// TIA Portal project "1215C_BREAKOUT_BOARD" (V19) (continued)
REGION Network 3
   RUNG wire#powerrail
      "FC10029_Custom_LGF_DTLtoString"(inDTL := "DB002-DateTime".LOCAL_DTL, format := 1, Ret_Val => "DB002-DateTime".DTLtoString_Ret, outDate_YY => "DB002-DateTime".sCustomDate_YY, outDate_MM => "DB002-DateTime".sCustomDate_MM, outDate_DD => "DB002-DateTime".sCustomDate_DD, outTime_HH => "DB002-DateTime".sCustomTime_HH, outTime_MM => "DB002-DateTime".sCustomTime_MM)
      "FC10030_Custom_DateTime_Format"(LOCAL_DTL := "DB002-DateTime".LOCAL_DTL, sCustomDate_YY := "DB002-DateTime".sCustomDate_YY, sCustomDate_MM := "DB002-DateTime".sCustomDate_MM, sCustomDate_DD := "DB002-DateTime".sCustomDate_DD, sCustomTime_HH := "DB002-DateTime".sCustomTime_HH, sCustomTime_MM := "DB002-DateTime".sCustomTime_MM, sCustomDate_DDMMYY := "DB002-DateTime".sCustomDate_DDMMYY, sCustomTime_HHMM := "DB002-DateTime".sCustomTime_HHMM)
   END_RUNG
   // the same network as SCL:
   "DB002-DateTime".DTLtoString_Ret := "FC10029_Custom_LGF_DTLtoString"(inDTL := "DB002-DateTime".LOCAL_DTL,
                           format := 1,
                           outDate_YY => "DB002-DateTime".sCustomDate_YY,
                           outDate_MM => "DB002-DateTime".sCustomDate_MM,
                           outDate_DD => "DB002-DateTime".sCustomDate_DD,
                           outTime_HH => "DB002-DateTime".sCustomTime_HH,
                           outTime_MM => "DB002-DateTime".sCustomTime_MM,
                           ENO => #_w1);
   IF #_w1 THEN
       "FC10030_Custom_DateTime_Format"(LOCAL_DTL := "DB002-DateTime".LOCAL_DTL,
                               sCustomDate_YY := "DB002-DateTime".sCustomDate_YY,
                               sCustomDate_MM := "DB002-DateTime".sCustomDate_MM,
                               sCustomDate_DD := "DB002-DateTime".sCustomDate_DD,
                               sCustomTime_HH := "DB002-DateTime".sCustomTime_HH,
                               sCustomTime_MM := "DB002-DateTime".sCustomTime_MM,
                               sCustomDate_DDMMYY := "DB002-DateTime".sCustomDate_DDMMYY,
                               sCustomTime_HHMM := "DB002-DateTime".sCustomTime_HHMM);
   END_IF;
END_REGION
END_FUNCTION

FUNCTION "FC10029_Custom_LGF_DTLtoString" : String   // FC10029, SCL
{ S7_Optimized_Access := 'TRUE' }
VERSION : 0.1
   VAR_INPUT
      inDTL : DTL;   // Date as DTL tag
      format : Bool;   // 1 = traditional, 0 = international
   END_VAR
   VAR_OUTPUT
      outDate_YY : String;   // Custom Date Output (YY)
      outDate_MM : String;   // Custom Date Output (MM)
      outDate_DD : String;   // Custom Date Output (DD)
      outTime_HH : String;   // Custom Time Output (HH)
      outTime_MM : String;   // Custom Time Output (MM)
   END_VAR
   VAR_TEMP
      tempString : String;   // -
      tempSepTime : Char;   // -
      tempPosYear : USInt;   // -
      tempPosMonth : USInt;   // -
      tempPosDay : USInt;   // -
      tempPosHour : USInt;   // -
      tempPosMinute : USInt;   // -
      tempPosSepYearMonth : USInt;   // -
      tempPosSepMonthDay : USInt;   // -
      tempPosSepHourMinute : USInt;   // -
   END_VAR
   // Ret_Val : Date as String tag
BEGIN
   //=============================================================================
   // Siemens AG
   // (c)Copyright 2017
   //-----------------------------------------------------------------------------
   // Library:       LGF (Library General Functions)
   // Tested with:   CPU1212C DC/DC/DC FW:V4.2
   // Engineering:   TIA Portal V14 Update 1
   // Restrictions:  -
   // Requirements:  PLC (S7-1200 / S7-1500)
   // Functionality: This function converts DTL into a string.  (EDITED)
   //-----------------------------------------------------------------------------
   // Change log table:
   // Version  Date        In charge / Changes applied
   // 01.00.00 15.06.2016  Siemens Industry Online Support
   //                      First released version
   // 01.00.01 02.01.2017  Siemens Industry Online Support
   //                      Upgrade: TIA Portal V14 Update 1
   // 01.00.02 17.08.2018  Siemens Industry Online Support
   //                      Upgrade: TIA V15 Update 2
   //=============================================================================


   // Initialization
   #tempString := '';
   #tempSepTime := ':';


   // Set format parameters for output string
   IF NOT #format
   THEN                                          // International ISO 8601
       #tempPosYear := 1;                          // DTL  | Y| Y| Y| Y| -| M| M| -| D| D|  | H| H| :| M| M|
       #tempPosMonth := 6;                         // -----|--|--|--|--|--|--|--|--|--|--|--|--|--|--|--|--|
       #tempPosDay := 9;                           // Pos  | 1| 2| 3| 4| 5| 6| 7| 8| 9|10|11|12|13|14|15|16|
       #tempPosHour := 12;
       #tempPosMinute := 15;
       #tempPosSepYearMonth := 5;
       #tempPosSepMonthDay := 8;
       #tempPosSepHourMinute := 14;
   ELSE                                          // Traditional (EU)
       #tempPosYear := 7;                          // DTL  | D| D| -| M| M| -| Y| Y| Y| Y|  | H| H| :| M| M|
       #tempPosMonth := 4;                         // -----|--|--|--|--|--|--|--|--|--|--|--|--|--|--|--|--|
       #tempPosDay := 1;                           // Pos  | 1| 2| 3| 4| 5| 6| 7| 8| 9|10|11|12|13|14|15|16|
       #tempPosHour := 12;
       #tempPosMinute := 15;
       #tempPosSepYearMonth := 6;
       #tempPosSepMonthDay := 3;
       #tempPosSepHourMinute := 14;
   END_IF;


   // Convert "Value" into "String" and place at the right position

   // Convert for YEAR
   VAL_STRG(FORMAT := W#16#0000,
            IN := #inDTL.YEAR,
            P := #tempPosYear,
            PREC := 0,
            SIZE := 4,
            OUT => #tempString);     // DTL YEAR --> String --> #tempPosYear

   VAL_STRG(FORMAT := W#16#0000,
            IN := #inDTL.YEAR MOD 100,
            P := 1,
            PREC := 0,
            SIZE := 2,
            OUT => #outDate_YY);        // DTL YEAR --> String --> #CustOutYear (Last 2 digits)

   // Convert for MONTH
   VAL_STRG(FORMAT := W#16#0000,
            IN := #inDTL.MONTH,
            P := #tempPosMonth,
            PREC := 0,
            SIZE := 2,
            OUT => #tempString);     // DTL MONTH --> String --> #tempPosMonth

   VAL_STRG(FORMAT := W#16#0000,
            IN := #inDTL.MONTH,
            P := 1,
            PREC := 0,
            SIZE := 2,
            OUT => #outDate_MM);        // DTL MONTH --> String --> #CustOutDate MM

   // Convert for DAY
   VAL_STRG(FORMAT := W#16#0000,
            IN := #inDTL.DAY,
            P := #tempPosDay,
            PREC := 0,
            SIZE := 2,
            OUT => #tempString);     // DTL DAY --> String --> #tempPosDay

   VAL_STRG(FORMAT := W#16#0000,
            IN := #inDTL.DAY,
            P := 1,
            PREC := 0,
            SIZE := 2,
            OUT => #outDate_DD);        // DTL DAY --> String --> #CustOutDate DDMM

   // Convert for HOUR
   VAL_STRG(FORMAT := W#16#0000,
            IN := #inDTL.HOUR,
            P := #tempPosHour,
            PREC := 0,
            SIZE := 2,
            OUT => #tempString);     // DTL HOUR --> String --> #tempPosHour

   VAL_STRG(FORMAT := W#16#0000,
            IN := #inDTL.HOUR,
            P := 1,
            PREC := 0,
            SIZE := 2,
            OUT => #outTime_HH);     // DTL HOUR --> String --> #CustOutTime HH

   // Convert for MINUTE
   VAL_STRG(FORMAT := W#16#0000,
            IN := #inDTL.MINUTE,
            P := #tempPosMinute,
            PREC := 0,
            SIZE := 2,
            OUT => #tempString);     // DTL MINUTE --> String --> #tempPosMinute

   VAL_STRG(FORMAT := W#16#0000,
            IN := #inDTL.MINUTE,
            P := 1,
            PREC := 0,
            SIZE := 2,
            OUT => #outTime_MM);        // DTL MINUTE --> String --> #CustOutTime


   // Block output
   #FC10029_Custom_LGF_DTLtoString := #tempString;


   // Additional outputs
   #outDate_YY := #outDate_YY;
   #outDate_MM := #outDate_MM;
   #outDate_DD := #outDate_DD;
   #outTime_HH := #outTime_HH;
   #outTime_MM := #outTime_MM;
END_FUNCTION

FUNCTION "FC10030_Custom_DateTime_Format" : Void   // FC10030, LAD
TITLE = Custom Date / Time Formats
{ S7_Optimized_Access := 'TRUE' }
VERSION : 0.1
   VAR_INPUT
      LOCAL_DTL : DTL;   // RAW DTL
   END_VAR
   VAR_IN_OUT
      sCustomDate_YY : String;   // Custom Year Output (YY)
      sCustomDate_MM : String;   // Custom Date Output (MM)
      sCustomDate_DD : String;   // Custom Date Output (DD)
      sCustomTime_HH : String;   // Custom Time Output (HH)
      sCustomTime_MM : String;   // Custom Time Output (MM)
      sCustomDate_DDMMYY : String;   // Custom Date (DD/MM/YY)
      sCustomTime_HHMM : String;   // Custom Date (HH:MM)
   END_VAR
   VAR_TEMP
      sTemp_String : String;   // -
   END_VAR
BEGIN

REGION Network 1: =================ADD_LEADING_ZEROS=================
END_REGION

REGION Network 2: Add leading zero to MM if less than 10
   // > If DTL.MONTH is less than 10 - replace 1st character in DD with a 0
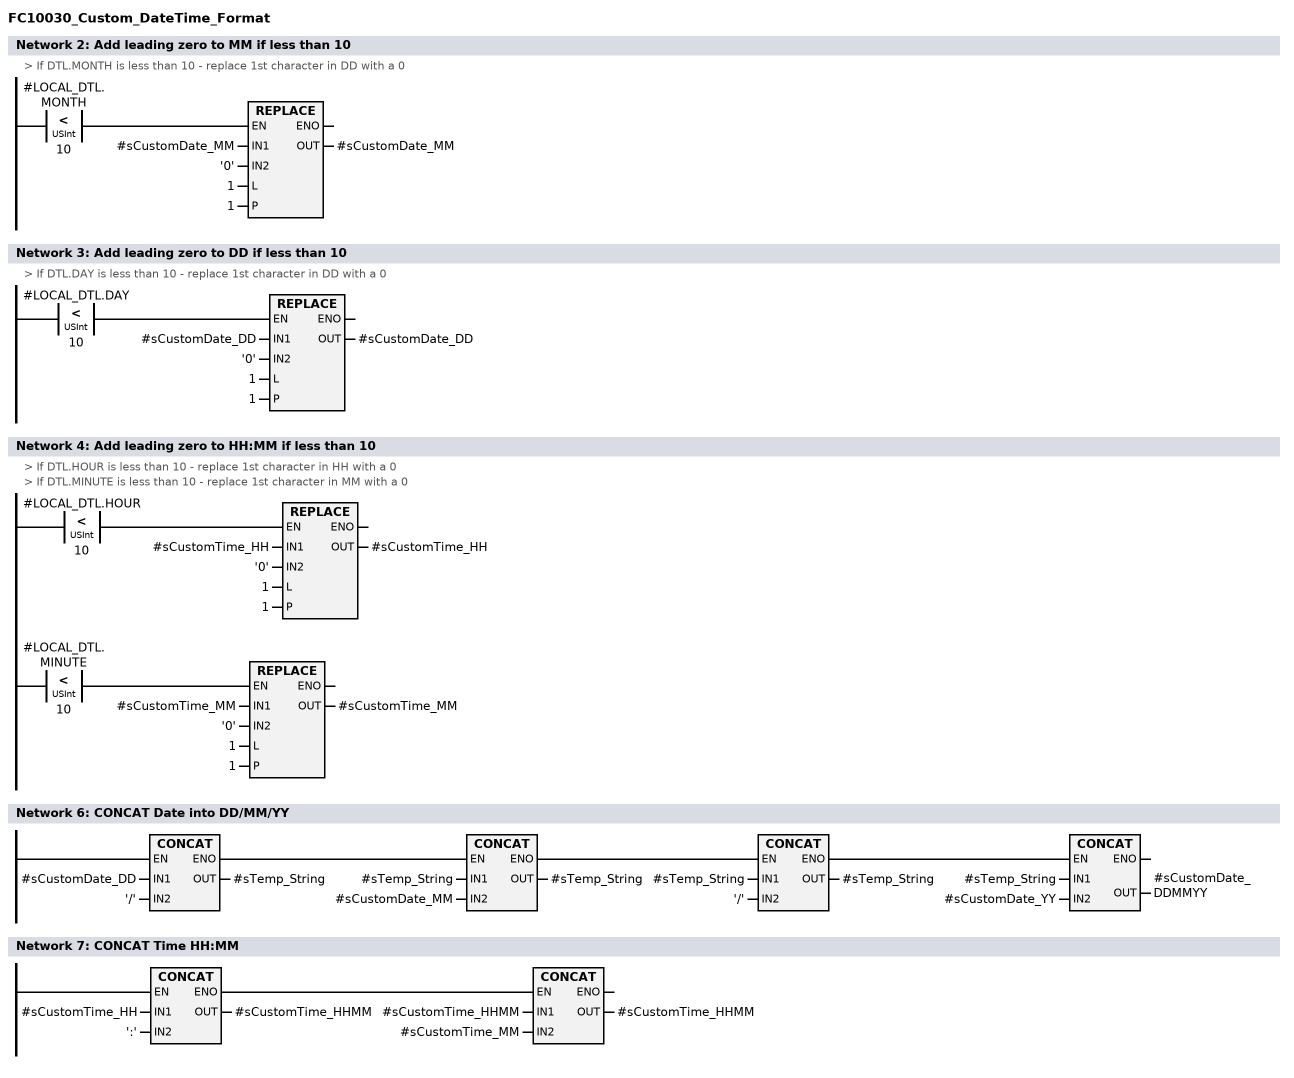
   IF #LOCAL_DTL.MONTH < 10 THEN
       #sCustomDate_MM := REPLACE(IN1 := #sCustomDate_MM, IN2 := '0', L := 1, P := 1);
   END_IF;
END_REGION

REGION Network 3: Add leading zero to DD if less than 10
   // > If DTL.DAY is less than 10 - replace 1st character in DD with a 0
   IF #LOCAL_DTL.DAY < 10 THEN
       #sCustomDate_DD := REPLACE(IN1 := #sCustomDate_DD, IN2 := '0', L := 1, P := 1);
   END_IF;
END_REGION

REGION Network 4: Add leading zero to HH:MM if less than 10
   // > If DTL.HOUR is less than 10 - replace 1st character in HH with a 0
   // > If DTL.MINUTE is less than 10 - replace 1st character in MM with a 0
   IF #LOCAL_DTL.HOUR < 10 THEN
       #sCustomTime_HH := REPLACE(IN1 := #sCustomTime_HH, IN2 := '0', L := 1, P := 1);
   END_IF;
   IF #LOCAL_DTL.MINUTE < 10 THEN
       #sCustomTime_MM := REPLACE(IN1 := #sCustomTime_MM, IN2 := '0', L := 1, P := 1);
   END_IF;
END_REGION

REGION Network 5: =================CONCAT_INTO_FORMAT=================
END_REGION

REGION Network 6: CONCAT Date into DD/MM/YY
   #sTemp_String := CONCAT(IN1 := #sCustomDate_DD, IN2 := '/');
   #sTemp_String := CONCAT(IN1 := #sTemp_String, IN2 := #sCustomDate_MM);
   #sTemp_String := CONCAT(IN1 := #sTemp_String, IN2 := '/');
   #sCustomDate_DDMMYY := CONCAT(IN1 := #sTemp_String, IN2 := #sCustomDate_YY);
END_REGION

REGION Network 7: CONCAT Time HH:MM
   #sCustomTime_HHMM := CONCAT(IN1 := #sCustomTime_HH, IN2 := ':');
   #sCustomTime_HHMM := CONCAT(IN1 := #sCustomTime_HHMM, IN2 := #sCustomTime_MM);
END_REGION
END_FUNCTION

(* ===== HMI "HMI_RT_1" =====
system functions are stored by id; their names below are inferred from use
connection "HMI_Connection": ETHERNET, SMART_S7_1200_OMS

HMI tags "Default tag table"
   "ScreenNumber" : UInt, internal

HMI tags "PLC_Inputs"
   "DB001-PLC_I/O_Inputs_xDI0.0" : Bool = PLC "DB001-PLC_I/O".Inputs."xDI0.0", 100 ms
   "DB001-PLC_I/O_Inputs_xDI0.1" : Bool = PLC "DB001-PLC_I/O".Inputs."xDI0.1", 100 ms
   "DB001-PLC_I/O_Inputs_xDI0.2" : Bool = PLC "DB001-PLC_I/O".Inputs."xDI0.2", 100 ms
   "DB001-PLC_I/O_Inputs_xDI0.3" : Bool = PLC "DB001-PLC_I/O".Inputs."xDI0.3", 100 ms
   "DB001-PLC_I/O_Inputs_xDI0.4" : Bool = PLC "DB001-PLC_I/O".Inputs."xDI0.4", 100 ms
   "DB001-PLC_I/O_Inputs_xDI0.5" : Bool = PLC "DB001-PLC_I/O".Inputs."xDI0.5", 100 ms
   "DB001-PLC_I/O_Inputs_xDI0.6" : Bool = PLC "DB001-PLC_I/O".Inputs."xDI0.6", 100 ms
   "DB001-PLC_I/O_Inputs_xDI0.7" : Bool = PLC "DB001-PLC_I/O".Inputs."xDI0.7", 100 ms
   "DB001-PLC_I/O_Inputs_xDI1.0" : Bool = PLC "DB001-PLC_I/O".Inputs."xDI1.0", 100 ms
   "DB001-PLC_I/O_Inputs_xDI1.1" : Bool = PLC "DB001-PLC_I/O".Inputs."xDI1.1", 100 ms
   "DB001-PLC_I/O_Inputs_xDI1.2" : Bool = PLC "DB001-PLC_I/O".Inputs."xDI1.2", 100 ms
   "DB001-PLC_I/O_Inputs_xDI1.3" : Bool = PLC "DB001-PLC_I/O".Inputs."xDI1.3", 100 ms
   "DB001-PLC_I/O_Inputs_xDI1.4" : Bool = PLC "DB001-PLC_I/O".Inputs."xDI1.4", 100 ms
   "DB001-PLC_I/O_Inputs_xDI1.5" : Bool = PLC "DB001-PLC_I/O".Inputs."xDI1.5", 100 ms

HMI tags "PLC_Outputs"
   "DB001-PLC_I/O_Outputs_xDQ0.0" : Bool = PLC "DB001-PLC_I/O".Outputs."xDQ0.0", 100 ms
   "DB001-PLC_I/O_Outputs_xDQ0.1" : Bool = PLC "DB001-PLC_I/O".Outputs."xDQ0.1", 100 ms
   "DB001-PLC_I/O_Outputs_xDQ0.2" : Bool = PLC "DB001-PLC_I/O".Outputs."xDQ0.2", 100 ms
   "DB001-PLC_I/O_Outputs_xDQ0.3" : Bool = PLC "DB001-PLC_I/O".Outputs."xDQ0.3", 100 ms
   "DB001-PLC_I/O_Outputs_xDQ0.4" : Bool = PLC "DB001-PLC_I/O".Outputs."xDQ0.4", 100 ms
   "DB001-PLC_I/O_Outputs_xDQ0.5" : Bool = PLC "DB001-PLC_I/O".Outputs."xDQ0.5", 100 ms
   "DB001-PLC_I/O_Outputs_xDQ0.6" : Bool = PLC "DB001-PLC_I/O".Outputs."xDQ0.6", 100 ms
   "DB001-PLC_I/O_Outputs_xDQ0.7" : Bool = PLC "DB001-PLC_I/O".Outputs."xDQ0.7", 100 ms
   "DB001-PLC_I/O_Outputs_xDQ1.0" : Bool = PLC "DB001-PLC_I/O".Outputs."xDQ1.0", 100 ms
   "DB001-PLC_I/O_Outputs_xDQ1.1" : Bool = PLC "DB001-PLC_I/O".Outputs."xDQ1.1", 100 ms

HMI tags "PLC_Analog"
   "AI0.0" : Word = PLC "AI0.0" AT %IW64, 100 ms
   "AQ0.0" : Word = PLC "AQ0.0" AT %QW64, 100 ms
   "DB001-PLC_I/O_Outputs_rAQ0.0_Scaled" : Real = PLC "DB001-PLC_I/O".Outputs."rAQ0.0_Scaled", 100 ms
   "DB001-PLC_I/O_Outputs_rAQ0.1_Scaled" : Real = PLC "DB001-PLC_I/O".Outputs."rAQ0.1_Scaled", 100 ms
   "AI0.1" : Word = PLC "AI0.1" AT %IW66, 100 ms
   "AQ0.1" : Word = PLC "AQ0.1" AT %QW66, 100 ms
   "DB001-PLC_I/O_Inputs_rAI0.0_Scaled" : Real = PLC "DB001-PLC_I/O".Inputs."rAI0.0_Scaled", 100 ms
   "DB001-PLC_I/O_Inputs_rAI0.1_Scaled" : Real = PLC "DB001-PLC_I/O".Inputs."rAI0.1_Scaled", 100 ms

HMI tags "PLC_DateTime"
   "DB002-DateTime_sCustomDate_DDMMYY" : String[254] = PLC "DB002-DateTime".sCustomDate_DDMMYY, 1 s
   "DB002-DateTime_sCustomTime_HHMM" : String[254] = PLC "DB002-DateTime".sCustomTime_HHMM, 1 s

text list "ON/OFF": 0 'OFF'; 1 'ON'

screen "01-Home" 480x272, template "Main_Template"
   on GenerateScreen: SetTag("ScreenNumber", 1)
   TextField "TextField_ProjectName" at 109,47 size 259x30; Text 'PLC BREAKOUT BOARD'
   TextField "Text field_DeviceInfo" at 21,91 size 435x52; Text '1215C DC/DC/DC -- 6ES7215-1AG40-0XB0 -- IP: 192.168.0.175/24 KTP400 HMI -- 6AV2123-2DB03-0AX0 -- IP: 192.168.0.176/24'
   TextField "Text field_Description" at 62,155 size 353x52; Text '- Displays the Digital & Analog Input states, - Toggle Digital Outputs via HMI buttons, - Simulation of Analog Outputs via 20 step incriments.'
   Button "Button_ExitRuntime" at 384,227 size 92x40; TextOff 'EXIT RUNTIME'
      on Press: StopRuntime(0)

screen "02-Inputs1" 480x272, template "Main_Template"
   on GenerateScreen: SetTag("ScreenNumber", 2)
   TextField "TextField_ScreenName" at 85,46 size 309x30; Text 'PLC DIGITAL INPUTS - 1of2'
   TextField "TextField_BankLetter" at 412,50 size 64x23; Text 'BANK A'
   Button "Button_Next" at 384,227 size 92x40; TextOff 'NEXT'
      on Press: ActivateScreen("03-Inputs2", 0)
   Group "Group_DI0.0" at 41,81 size 62x63
   Group "Group_DI0.1" at 153,81 size 62x63
   Group "Group_DI0.2" at 265,81 size 62x63
   Group "Group_DI0.3" at 377,81 size 62x63
   Group "Group_DI0.4" at 41,152 size 62x64
   Group "Group_DI0.5" at 153,152 size 62x64
   Group "Group_DI0.6" at 265,154 size 62x64
   Group "Group_DI0.7" at 377,154 size 62x64
   TextField "Text field_DI0.0" at 51,81 size 42x19; Text 'DI 0.0'
   Circle "Circle_DI0.0" at 54,103 size 36x36
      Appearance <- "DB001-PLC_I/O_Inputs_xDI0.0"
   TextField "Text field_DI0.1" at 163,81 size 42x19; Text 'DI 0.1'
   Circle "Circle_DI0.1" at 166,103 size 36x36
      Appearance <- "DB001-PLC_I/O_Inputs_xDI0.1"
   TextField "Text field_DI0.2" at 275,81 size 42x19; Text 'DI 0.2'
   Circle "Circle_DI0.2" at 278,103 size 36x36
      Appearance <- "DB001-PLC_I/O_Inputs_xDI0.2"
   TextField "Text field_DI0.3" at 387,81 size 42x19; Text 'DI 0.3'
   Circle "Circle_DI0.3" at 390,103 size 36x36
      Appearance <- "DB001-PLC_I/O_Inputs_xDI0.3"
   TextField "Text field_DI0.4" at 51,152 size 42x19; Text 'DI 0.4'
   Circle "Circle_DI0.4" at 54,174 size 36x36
      Appearance <- "DB001-PLC_I/O_Inputs_xDI0.4"
   TextField "Text field_DI0.5" at 163,152 size 42x19; Text 'DI 0.5'
   Circle "Circle_DI0.5" at 166,174 size 36x36
      Appearance <- "DB001-PLC_I/O_Inputs_xDI0.5"
   TextField "Text field_DI0.6" at 275,154 size 42x19; Text 'DI 0.6'
   Circle "Circle_DI0.6" at 278,176 size 36x36
      Appearance <- "DB001-PLC_I/O_Inputs_xDI0.6"
   TextField "Text field_DI0.7" at 387,154 size 42x19; Text 'DI 0.7'
   Circle "Circle_DI0.7" at 390,176 size 36x36
      Appearance <- "DB001-PLC_I/O_Inputs_xDI0.7"

screen "04-Outputs1" 480x272, template "Main_Template"
   on GenerateScreen: SetTag("ScreenNumber", 4)
   TextField "TextField_ScreenName" at 76,46 size 328x30; Text 'PLC DIGITAL OUTPUTS - 1of2'
   TextField "TextField_BankLetter" at 412,50 size 64x23; Text 'BANK A'
   Button "Button_Next" at 384,227 size 92x40; TextOff 'NEXT'
      on Press: ActivateScreen("05-Outputs2", 0)
   Group "Group_DQ0.0" at 18,83 size 97x62; TextList "ON/OFF"
   Group "Group_DQ0.1" at 132,83 size 97x62; TextList "ON/OFF"
   Group "Group_DQ0.2" at 247,83 size 97x62; TextList "ON/OFF"
   Group "Group_DQ0.3" at 362,83 size 97x62; TextList "ON/OFF"
   Group "Group_DQ0.4" at 18,154 size 97x62; TextList "ON/OFF"
   Group "Group_DQ0.5" at 132,154 size 97x62; TextList "ON/OFF"
   Group "Group_DQ0.6" at 247,154 size 97x62; TextList "ON/OFF"
   Group "Group_DQ0.7" at 362,154 size 97x62; TextList "ON/OFF"
   Rectangle "Rectangle_DQ0.0" at 18,83 size 97x62
      Appearance <- "DB001-PLC_I/O_Outputs_xDQ0.0"
   TextField "Text field_DQ0.0" at 44,83 size 46x19; Text 'DQ 0.0'
   Button "Button_DQ0.0" at 30,105 size 73x32; TextOff 'Text'; TextList "ON/OFF"
      on Press: InvertBit("DB001-PLC_I/O_Outputs_xDQ0.0")
      ProcessValue <- "DB001-PLC_I/O_Outputs_xDQ0.0"
   Rectangle "Rectangle_DQ0.1" at 132,83 size 97x62
      Appearance <- "DB001-PLC_I/O_Outputs_xDQ0.1"
   TextField "Text field_DQ0.1" at 158,83 size 46x19; Text 'DQ 0.1'
   Button "Button_DQ0.1" at 144,105 size 73x32; TextOff 'Text'; TextList "ON/OFF"
      on Press: InvertBit("DB001-PLC_I/O_Outputs_xDQ0.1")
      ProcessValue <- "DB001-PLC_I/O_Outputs_xDQ0.1"
   Rectangle "Rectangle_DQ0.2" at 247,83 size 97x62
      Appearance <- "DB001-PLC_I/O_Outputs_xDQ0.2"
   TextField "Text field_DQ0.2" at 273,83 size 46x19; Text 'DQ 0.2'
   Button "Button_DQ0.2" at 259,105 size 73x32; TextOff 'Text'; TextList "ON/OFF"
      on Press: InvertBit("DB001-PLC_I/O_Outputs_xDQ0.2")
      ProcessValue <- "DB001-PLC_I/O_Outputs_xDQ0.2"
   Rectangle "Rectangle_DQ0.3" at 362,83 size 97x62
      Appearance <- "DB001-PLC_I/O_Outputs_xDQ0.3"
   TextField "Text field_DQ0.3" at 388,83 size 46x19; Text 'DQ 0.3'
   Button "Button_DQ0.3" at 374,105 size 73x32; TextOff 'Text'; TextList "ON/OFF"
      on Press: InvertBit("DB001-PLC_I/O_Outputs_xDQ0.3")
      ProcessValue <- "DB001-PLC_I/O_Outputs_xDQ0.3"
   Rectangle "Rectangle_DQ0.4" at 18,154 size 97x62
      Appearance <- "DB001-PLC_I/O_Outputs_xDQ0.4"
   TextField "Text field_DQ0.4" at 44,154 size 46x19; Text 'DQ 0.4'
   Button "Button_DQ0.4" at 30,176 size 73x32; TextOff 'Text'; TextList "ON/OFF"
      on Press: InvertBit("DB001-PLC_I/O_Outputs_xDQ0.4")
      ProcessValue <- "DB001-PLC_I/O_Outputs_xDQ0.4"
   Rectangle "Rectangle_DQ0.5" at 132,154 size 97x62
      Appearance <- "DB001-PLC_I/O_Outputs_xDQ0.5"
   TextField "Text field_DQ0.5" at 158,154 size 46x19; Text 'DQ 0.5'
   Button "Button_DQ0.5" at 144,176 size 73x32; TextOff 'Text'; TextList "ON/OFF"
      on Press: InvertBit("DB001-PLC_I/O_Outputs_xDQ0.5")
      ProcessValue <- "DB001-PLC_I/O_Outputs_xDQ0.5"
   Rectangle "Rectangle_DQ0.6" at 247,154 size 97x62
      Appearance <- "DB001-PLC_I/O_Outputs_xDQ0.6"
   TextField "Text field_DQ0.6" at 273,154 size 46x19; Text 'DQ 0.6'
   Button "Button_DQ0.6" at 259,176 size 73x32; TextOff 'Text'; TextList "ON/OFF"
      on Press: InvertBit("DB001-PLC_I/O_Outputs_xDQ0.6")
      ProcessValue <- "DB001-PLC_I/O_Outputs_xDQ0.6"
   Rectangle "Rectangle_DQ0.7" at 362,154 size 97x62
      Appearance <- "DB001-PLC_I/O_Outputs_xDQ0.7"
   TextField "Text field_DQ0.7" at 388,154 size 46x19; Text 'DQ 0.7'
   Button "Button_DQ0.7" at 374,176 size 73x32; TextOff 'Text'; TextList "ON/OFF"
      on Press: InvertBit("DB001-PLC_I/O_Outputs_xDQ0.7")
      ProcessValue <- "DB001-PLC_I/O_Outputs_xDQ0.7"

screen "06-AnalogI/O" 480x272, template "Main_Template"
   on GenerateScreen: SetTag("ScreenNumber", 6)
   Button "Button_Back" at 384,227 size 92x40; TextOff 'BACK'
      on Press: function_efd93a16()
   TextField "TextField_ScreenName" at 65,46 size 351x30; Text 'PLC ANALOG INPUTS/OUTPUTS'
   Group "Group_A0" at 244,76 size 229x145; FormatPattern 9999
   Group "Group_A1" at 8,76 size 229x145; FormatPattern 9999
   TextField "Text field_A0" at 291,77 size 127x21; Text 'Analog AI-0 & AQ-0'
   TextField "Text field_A0_Input" at 279,98 size 42x17; Text 'INPUT'
   TextField "Text field_A0_Instruction" at 256,115 size 86x34; Text 'Use the connected potentiometer to change the input voltage.'
   TextField "Text field_A0_Voltage" at 280,149 size 41x14; Text 'VOLTAGE:'
   IOField "I/O field_A0_Voltage" at 281,162 size 42x21; FormatPattern 99.99; Unit  V
      ProcessValue <- "DB001-PLC_I/O_Inputs_rAI0.0_Scaled"
   TextField "Text field_A0_InRAW" at 289,181 size 24x14; Text 'RAW:'
   IOField "I/O field_A0_RAW" at 283,193 size 37x21; FormatPattern 99999
      ProcessValue <- "AI0.0"
   TextField "Text field_A0_Output" at 389,98 size 52x17; Text 'OUTPUT'
   TextField "Text field_A0_mA" at 381,127 size 19x14; Text 'mA:'
   IOField "I/O field_A0_mA" at 365,140 size 51x21; FormatPattern 99.99; Unit  mA
      ProcessValue <- "DB001-PLC_I/O_Outputs_rAQ0.0_Scaled"
   TextField "Text field_A0_OutRAW" at 379,167 size 24x14; Text 'RAW:'
   IOField "I/O field_A0_OutRAW" at 373,180 size 37x21; FormatPattern 99999
      ProcessValue <- "AQ0.0"
   TextField "Text field_A0_20" at 403,113 size 25x14; Text '20mA'
   TextField "Text field_A0_15" at 415,136 size 13x14; Text '15'
   TextField "Text field_A0_10" at 415,160 size 13x14; Text '10'
   TextField "Text field_A0_5" at 419,182 size 10x14; Text '5'
   TextField "Text field_A0_0" at 408,205 size 21x14; Text '0mA'
   Bar "Bar_A0" at 428,118 size 37x97; MinimumValue 0; MaximumValue 20
      ProcessValue <- "DB001-PLC_I/O_Outputs_rAQ0.0_Scaled"
   TextField "Text field_A1" at 55,77 size 127x21; Text 'Analog AI-1 & AQ-1'
   TextField "Text field_A1_Input" at 43,98 size 42x17; Text 'INPUT'
   TextField "Text field_A1_Instruction" at 20,115 size 86x34; Text 'Use the connected potentiometer to change the input voltage.'
   TextField "Text field_A1_Voltage" at 44,149 size 41x14; Text 'VOLTAGE:'
   IOField "I/O field_A1_Voltage" at 45,162 size 42x21; FormatPattern 99.99; Unit  V
      ProcessValue <- "DB001-PLC_I/O_Inputs_rAI0.1_Scaled"
   TextField "Text field_A1_InRAW" at 53,181 size 24x14; Text 'RAW:'
   IOField "I/O field_A1_RAW" at 47,193 size 37x21; FormatPattern 99999
      ProcessValue <- "AI0.1"
   TextField "Text field_A1_Output" at 153,98 size 52x17; Text 'OUTPUT'
   TextField "Text field_A1_mA" at 145,127 size 19x14; Text 'mA:'
   IOField "I/O field_A1_mA" at 129,140 size 51x21; FormatPattern 99.99; Unit  mA
      ProcessValue <- "DB001-PLC_I/O_Outputs_rAQ0.1_Scaled"
   TextField "Text field_A1_OutRAW" at 143,167 size 24x14; Text 'RAW:'
   IOField "I/O field_A1_OutRAW" at 137,180 size 37x21; FormatPattern 99999
      ProcessValue <- "AQ0.1"
   TextField "Text field_A1_20" at 167,113 size 25x14; Text '20mA'
   TextField "Text field_A1_15" at 179,136 size 13x14; Text '15'
   TextField "Text field_A1_10" at 179,160 size 13x14; Text '10'
   TextField "Text field_A1_5" at 183,182 size 10x14; Text '5'
   TextField "Text field_A1_0" at 172,205 size 21x14; Text '0mA'
   Bar "Bar_A1" at 192,118 size 37x97; MinimumValue 0; MaximumValue 20
      ProcessValue <- "DB001-PLC_I/O_Outputs_rAQ0.1_Scaled"

screen "03-Inputs2" 480x272, template "Main_Template"
   on GenerateScreen: SetTag("ScreenNumber", 3)
   Button "Button_Back" at 384,227 size 92x40; TextOff 'BACK'
      on Press: function_efd93a16()
   TextField "TextField_ScreenName" at 85,46 size 309x30; Text 'PLC DIGITAL INPUTS - 2of2'
   TextField "TextField_BankLetter" at 412,50 size 62x23; Text 'BANK B'
   Group "Group_DI1.0" at 73,81 size 62x63
   Group "Group_DI1.1" at 209,81 size 62x63
   Group "Group_DI1.2" at 345,81 size 62x63
   Group "Group_DI1.3" at 73,152 size 62x63
   Group "Group_DI1.4" at 209,152 size 62x64
   Group "Group_DI1.5" at 345,152 size 62x64
   TextField "Text field_DI1.0" at 83,81 size 42x19; Text 'DI 1.0'
   Circle "Circle_DI1.0" at 86,103 size 36x36
      Appearance <- "DB001-PLC_I/O_Inputs_xDI1.0"
   TextField "Text field_DI1.1" at 219,81 size 42x19; Text 'DI 1.1'
   Circle "Circle_DI1.1" at 222,103 size 36x36
      Appearance <- "DB001-PLC_I/O_Inputs_xDI1.1"
   TextField "Text field_DI1.2" at 355,81 size 42x19; Text 'DI 1.2'
   Circle "Circle_DI1.2" at 358,103 size 36x36
      Appearance <- "DB001-PLC_I/O_Inputs_xDI1.2"
   TextField "Text field_DI1.3" at 83,152 size 42x19; Text 'DI 1.3'
   Circle "Circle_DI1.3" at 86,174 size 36x36
      Appearance <- "DB001-PLC_I/O_Inputs_xDI1.3"
   TextField "Text field_DI1.4" at 219,152 size 42x19; Text 'DI 1.4'
   Circle "Circle_DI1.4" at 222,174 size 36x36
      Appearance <- "DB001-PLC_I/O_Inputs_xDI1.4"
   TextField "Text field_DI1.5" at 355,152 size 42x19; Text 'DI 1.5'
   Circle "Circle_DI1.5" at 358,174 size 36x36
      Appearance <- "DB001-PLC_I/O_Inputs_xDI1.5"

screen "05-Outputs2" 480x272, template "Main_Template"
   on GenerateScreen: SetTag("ScreenNumber", 5)
   TextField "TextField_ScreenName" at 76,46 size 328x30; Text 'PLC DIGITAL OUTPUTS - 2of2'
   TextField "TextField_BankLetter" at 412,50 size 62x23; Text 'BANK B'
   Button "Button_Back" at 384,227 size 92x40; TextOff 'BACK'
      on Press: function_efd93a16()
   Rectangle "Rectangle_DQ1.0" at 119,114 size 97x62
      Appearance <- "DB001-PLC_I/O_Outputs_xDQ1.0"
   TextField "Text field_DQ1.0" at 145,114 size 46x19; Text 'DQ 1.0'
   Button "Button_DQ1.0" at 131,136 size 73x32; TextOff 'Text'; TextList "ON/OFF"
      on Press: InvertBit("DB001-PLC_I/O_Outputs_xDQ1.0")
      ProcessValue <- "DB001-PLC_I/O_Outputs_xDQ0.0"
   Group "Group_DQ1.0" at 119,114 size 97x62; TextList "ON/OFF"
   Group "Group_DQ1.1" at 264,114 size 97x62; TextList "ON/OFF"
   Rectangle "Rectangle_DQ1.1" at 264,114 size 97x62
      Appearance <- "DB001-PLC_I/O_Outputs_xDQ1.1"
   TextField "Text field_DQ1.1" at 290,114 size 46x19; Text 'DQ 1.1'
   Button "Button_DQ1.1" at 276,136 size 73x32; TextOff 'Text'; TextList "ON/OFF"
      on Press: InvertBit("DB001-PLC_I/O_Outputs_xDQ1.1")
      ProcessValue <- "DB001-PLC_I/O_Outputs_xDQ0.1"

Template "Main_Template" 480x272
   GraphicView "Template_Background" at 0,0 size 480x272; Picture "HMI_Background"
   Button "Template_Button5_Blank" at 384,227 size 92x40; TextOff 'BLANK'
   Button "Template_Button1_Home" at 4,227 size 92x40; TextOff 'HOME'
      on Press: ActivateScreen("01-Home", 0)
   Button "Template_Button2_Inputs" at 99,227 size 92x40; TextOff 'INPUTS'
      on Press: ActivateScreen("02-Inputs1", 0)
   Button "Template_Button3_Outputs" at 194,227 size 92x40; TextOff 'OUTPUTS'
      on Press: ActivateScreen("04-Outputs1", 0)
   Button "Template_Button4_AnalogIO" at 289,227 size 92x40; TextOff 'ANALOG I/O'
      on Press: ActivateScreen("06-AnalogI/O", 0)
   IOField "Template_I/O field_Date" at 289,14 size 74x20; FormatPattern ????????
      ProcessValue <- "DB002-DateTime_sCustomDate_DDMMYY"
   IOField "Template_I/O field_Time" at 365,14 size 50x20; FormatPattern ?????
      ProcessValue <- "DB002-DateTime_sCustomTime_HHMM"
   GraphicView "TVET_Logo" at 8,2 size 220x44; Picture "TVET_Logo"
*)